(* Logix 5000 project; controller MV vendor 1 type 14 code 217 rev 31.11; software revision 31.00; part 5 of 53 *)
(* tags used below, declared in another part *)
   Always_Off : BOOL;
   Always_On : BOOL;
   ChangeDayONS : BOOL;
   CheckTimeMask : INT;
   CLOCKsetvalues : DINT[7];
   CurrentTime : DateTime;
   CWD : CHECKWORD_FLAGS;
   FtoF_raw_input : REAL;
   ItoF_raw_input : INT;
   MC_ALARM_RETURNED_STRING : STRING;
   MC_CH1_Log_ID : DINT;
   MC_CH2_Log_ID : DINT;
   MC_Channel1_Channel_1_event : STRING;
   MC_Channel1_Channel_1_event_prefix : STRING;
   MC_Channel1_Channel_2_event : STRING;
   MC_Channel1_Channel_2_event_prefix : STRING;
   MC_CLOCK_system_set : BOOL;
   MC_DetTank1_Service_event : STRING;
   MC_DetTank1_Service_event_prefix : STRING;
   MC_DetTank2_Service_event : STRING;
   MC_DetTank2_Service_event_prefix : STRING;
   MC_Event_Alarm_Tag : ALARM_DIGITAL;
   MC_Event_control_FIFO : CONTROL;
   MC_Event_control_FIFO_Operation_Type : CONTROL;
   MC_Event_Delay_For_Data : TIMER;
   MC_Event_Delay_For_PLC_Startup_Data : TIMER;
   MC_Event_Delay_Timer : TIMER;
   MC_Event_Delay_Timer_Off : TIMER;
   MC_Event_from_buffer : STRING;
   MC_Event_from_buffer_LogData1 : REAL;
   MC_Event_from_buffer_LogData2 : REAL;
   MC_Event_from_buffer_LogData3 : REAL;
   MC_Event_from_buffer_LogData4 : REAL;
   MC_Event_from_buffer_Operation_Type : DINT;
   MC_event_step : DINT;
   MC_Event_String_Last : STRING;
   MC_Event_Transact_Trigger_Tag : DINT;
   MC_Events_FIFO_Buffer : STRING[31];
   MC_Events_FIFO_Buffer_Operation_Type : INT[31];
   MC_Last_LogData_For_Op : REAL[60,20];
   MC_N10 : INT[255];   // SETTINGS
   MC_N100 : INT[255];   // C1_PLC Channel 1 PLC data
   MC_N100_20_alarm : ALARM_DIGITAL;
   MC_N100_20_Alarm_Ready : BOOL;
   MC_N100_20_Delayed_Timer2 : TIMER;
   MC_N100_20_Fault_Returned : STRING;
   MC_N100_20_SQL_Done : DINT;
   MC_N100_23_alarm : ALARM_DIGITAL;
   MC_N100_23_Alarm_Ready : BOOL;
   MC_N100_23_Delayed_Timer2 : TIMER;
   MC_N100_23_Event_Returned : STRING;
   MC_N100_23_SQL_Done : DINT;
   MC_N120 : INT[255];   // C2 PLC Channel 2 PLC data
   MC_N120_20_alarm : ALARM_DIGITAL;
   MC_N120_20_Alarm_Ready : BOOL;
   MC_N120_20_Delayed_Timer2 : TIMER;
   MC_N120_20_Fault_Returned : STRING;
   MC_N120_20_SQL_Done : DINT;
   MC_N120_23_alarm : ALARM_DIGITAL;
   MC_N120_23_Alarm_Ready : BOOL;
   MC_N120_23_Delayed_Timer2 : TIMER;
   MC_N120_23_Event_Returned : STRING;
   MC_N120_23_SQL_Done : DINT;
   MC_N140 : INT[31];   // RT FILL RT filling routine d ata
   MC_N160 : INT[255];   // P40 CHECK
   MC_N80 : INT[255];   // SRV1_PLC Detergent tank 1 ser vice PLC data
   MC_N80_10_alarm : ALARM_DIGITAL;
   MC_N80_10_Alarm_Ready : BOOL;
   MC_N80_10_Delayed_Timer2 : TIMER;
   MC_N80_10_Fault_Returned : STRING;
   MC_N80_10_SQL_Done : DINT;
   MC_N80_13_alarm : ALARM_DIGITAL;
   MC_N80_13_Alarm_Ready : BOOL;
   MC_N80_13_Delayed_Timer2 : TIMER;
   MC_N80_13_Event_Returned : STRING;
   MC_N80_13_SQL_Done : DINT;
   MC_N90 : INT[255];   // SV2_PLC Detergent tank 2 ser vice PLC data
   MC_N90_10_alarm : ALARM_DIGITAL;
   MC_N90_10_Alarm_Ready : BOOL;
   MC_N90_10_Delayed_Timer2 : TIMER;
   MC_N90_10_Fault_Returned : STRING;
   MC_N90_10_SQL_Done : DINT;
   MC_N90_13_alarm : ALARM_DIGITAL;
   MC_N90_13_Alarm_Ready : BOOL;
   MC_N90_13_Delayed_Timer2 : TIMER;
   MC_N90_13_Event_Returned : STRING;
   MC_N90_13_SQL_Done : DINT;
   MC_RT_Emptying_Log_ID : DINT;
   MC_RT_Filling_Log_ID : DINT;
   MC_SFile : INT[255];   // SLC Equivalent System File, So Original Code Can Remain
   MC_SRV1_Log_ID : DINT;
   MC_SRV2_Log_ID : DINT;
   One_Minute_One_Scan : BOOL;
   One_Minute_One_Scan_Timer : TIMER;
   One_Second_1_scan : BOOL;
   One_Second_One_Scan : ALIAS FOR One_Second_1_scan;
   scada_watchdog : DINT;
   scale_analog_int : DINT;
   scale_analog_result : REAL;
   scale_eu_max : REAL;
   scale_eu_min : REAL;
   scale_raw_input : REAL;
   scale_raw_max : REAL;
   scale_raw_min : REAL;
   scale_routine_active : BOOL;
   scale_temp : REAL;
(* MC_Common, continued *)

ROUTINE Analog_scale_ftof   (* ladder *)
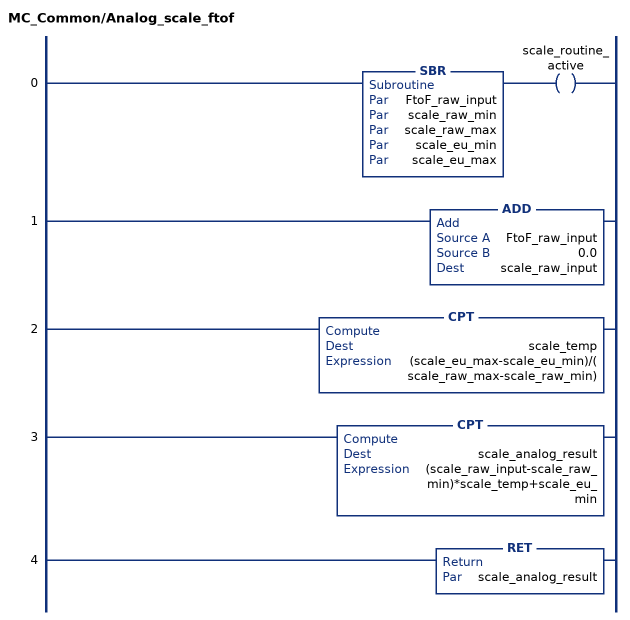
   0: SBR(FtoF_raw_input,scale_raw_min,scale_raw_max,scale_eu_min,scale_eu_max)OTE(scale_routine_active);
   1: ADD(FtoF_raw_input,0.0,scale_raw_input);
   2: CPT(scale_temp,(scale_eu_max-scale_eu_min)/(scale_raw_max-scale_raw_min));
   3: CPT(scale_analog_result,(scale_raw_input-scale_raw_min)*scale_temp+scale_eu_min);
   4: RET(scale_analog_result);
END_ROUTINE

ROUTINE Analog_Scale_FtoI   (* ladder *)
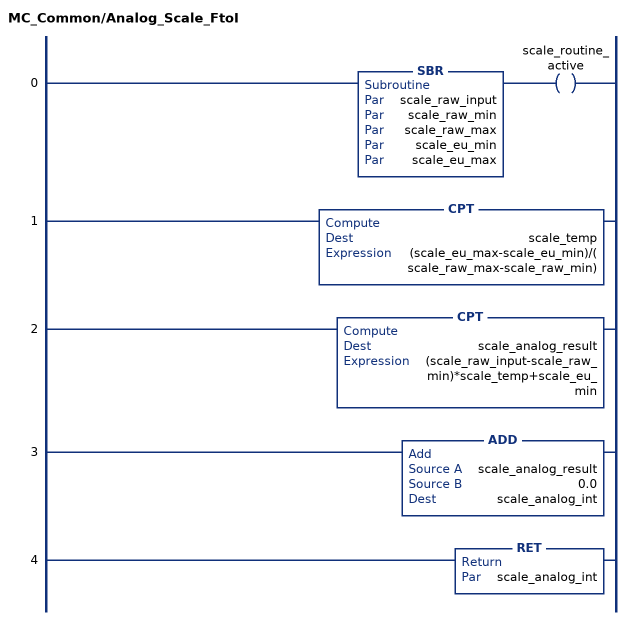
   0: SBR(scale_raw_input,scale_raw_min,scale_raw_max,scale_eu_min,scale_eu_max)OTE(scale_routine_active);
   1: CPT(scale_temp,(scale_eu_max-scale_eu_min)/(scale_raw_max-scale_raw_min));
   2: CPT(scale_analog_result,(scale_raw_input-scale_raw_min)*scale_temp+scale_eu_min);
   3: ADD(scale_analog_result,0.0,scale_analog_int);
   4: RET(scale_analog_int);
END_ROUTINE

ROUTINE Analog_Scale_ItoF   (* ladder *)
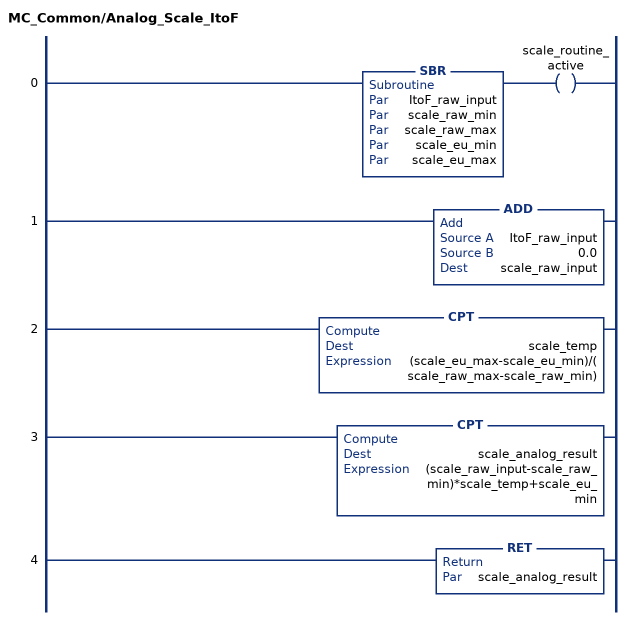
   0: SBR(ItoF_raw_input,scale_raw_min,scale_raw_max,scale_eu_min,scale_eu_max)OTE(scale_routine_active);
   1: ADD(ItoF_raw_input,0.0,scale_raw_input);
   2: CPT(scale_temp,(scale_eu_max-scale_eu_min)/(scale_raw_max-scale_raw_min));
   3: CPT(scale_analog_result,(scale_raw_input-scale_raw_min)*scale_temp+scale_eu_min);
   4: RET(scale_analog_result);
END_ROUTINE

ROUTINE ClockRoutines   (* ladder *)
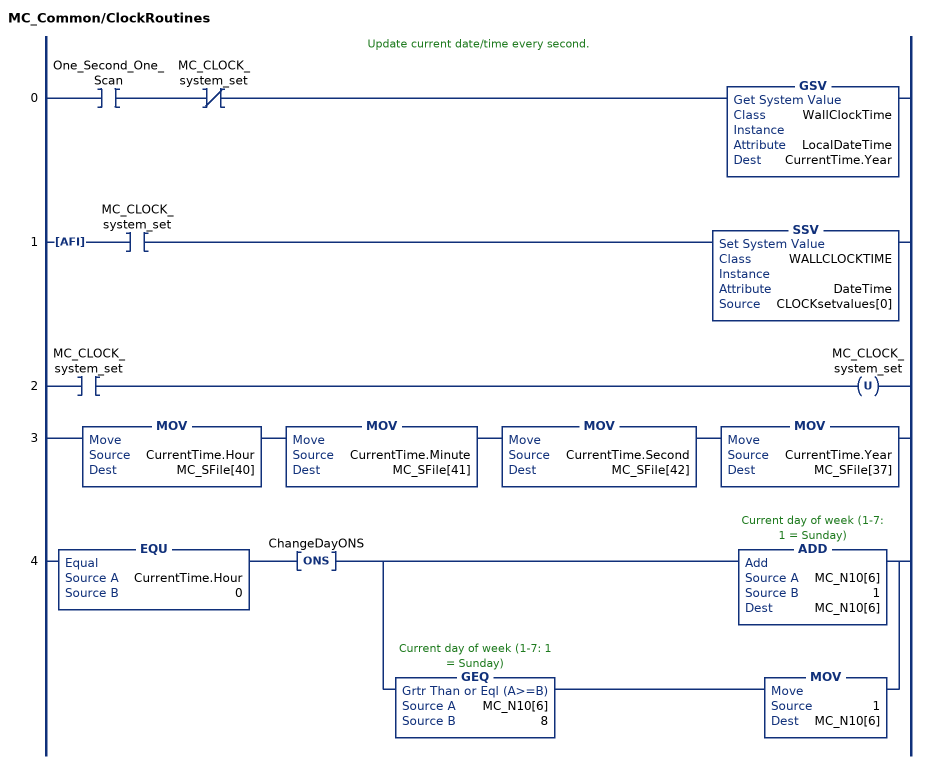
   // Update current date/time every second.
   0: XIC(One_Second_One_Scan)XIO(MC_CLOCK_system_set)GSV(WallClockTime,,LocalDateTime,CurrentTime.Year);
   1: AFI()XIC(MC_CLOCK_system_set)SSV(WALLCLOCKTIME,,DateTime,CLOCKsetvalues[0]);
   2: XIC(MC_CLOCK_system_set)OTU(MC_CLOCK_system_set);
   3: MOV(CurrentTime.Hour,MC_SFile[40])MOV(CurrentTime.Minute,MC_SFile[41])MOV(CurrentTime.Second,MC_SFile[42])MOV(CurrentTime.Year,MC_SFile[37]);
   4: EQU(CurrentTime.Hour,0)ONS(ChangeDayONS)[ADD(MC_N10[6],1,MC_N10[6]) ,GEQ(MC_N10[6],8) MOV(1,MC_N10[6]) ];
END_ROUTINE

ROUTINE Constants   (* ladder *)
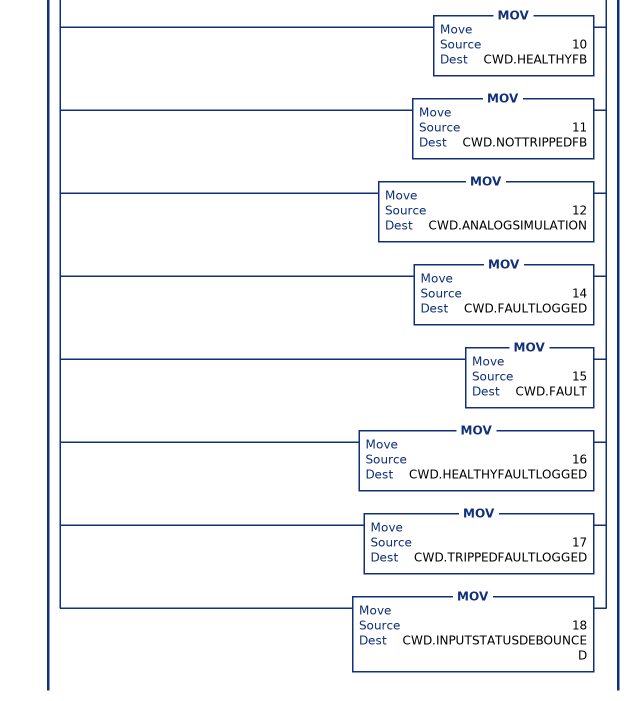
   0: [MOV(0,CWD.AUTODRV) ,MOV(0,CWD.INPUTSTATUS) ,MOV(1,CWD.PREVSCAN) ,MOV(2,CWD.SIMFAIL) ,MOV(3,CWD.OPENFB) ,MOV(3,CWD.RUNFB) ,MOV(4,CWD.CLOSEDFB) ,MOV(5,CWD.MANDRV) ,MOV(6,CWD.MANUAL) ,MOV(7,CWD.OUTPUT) ,MOV(8,CWD.CHECKOFF) ,MOV(9,CWD.HIGHLIGHT) ,MOV(10,CWD.HEALTHYFB) ,MOV(11,CWD.NOTTRIPPEDFB) ,MOV(12,CWD.ANALOGSIMULATION) ,MOV(14,CWD.FAULTLOGGED) ,MOV(15,CWD.FAULT) ,MOV(16,CWD.HEALTHYFAULTLOGGED) ,MOV(17,CWD.TRIPPEDFAULTLOGGED) ,MOV(18,CWD.INPUTSTATUSDEBOUNCED) ];
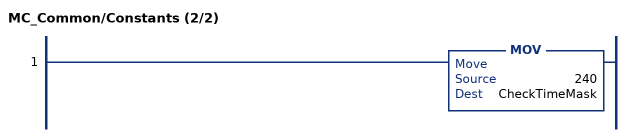
   1: MOV(240,CheckTimeMask);
END_ROUTINE

ROUTINE general_timers   (* ladder *)
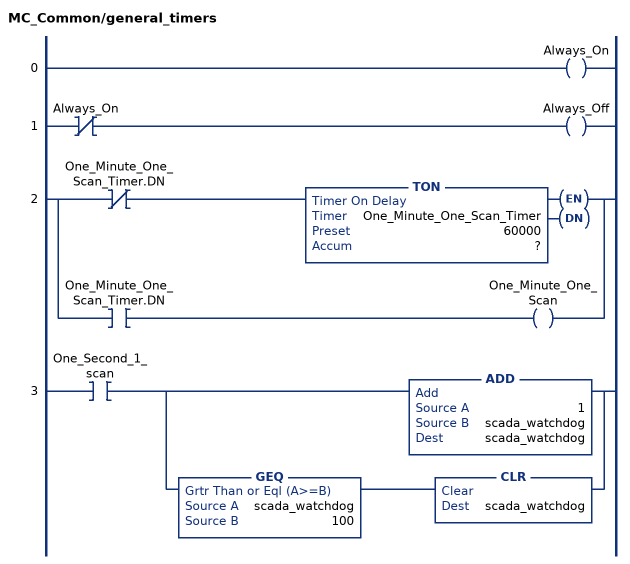
   0: OTE(Always_On);
   1: XIO(Always_On)OTE(Always_Off);
   2: [XIO(One_Minute_One_Scan_Timer.DN) TON(One_Minute_One_Scan_Timer,?,?) ,XIC(One_Minute_One_Scan_Timer.DN) OTE(One_Minute_One_Scan) ];
   3: XIC(One_Second_1_scan)[ADD(1,scada_watchdog,scada_watchdog) ,GEQ(scada_watchdog,100) CLR(scada_watchdog) ];
END_ROUTINE

ROUTINE MC_A_Alarms_From_PLC   (* ladder *)
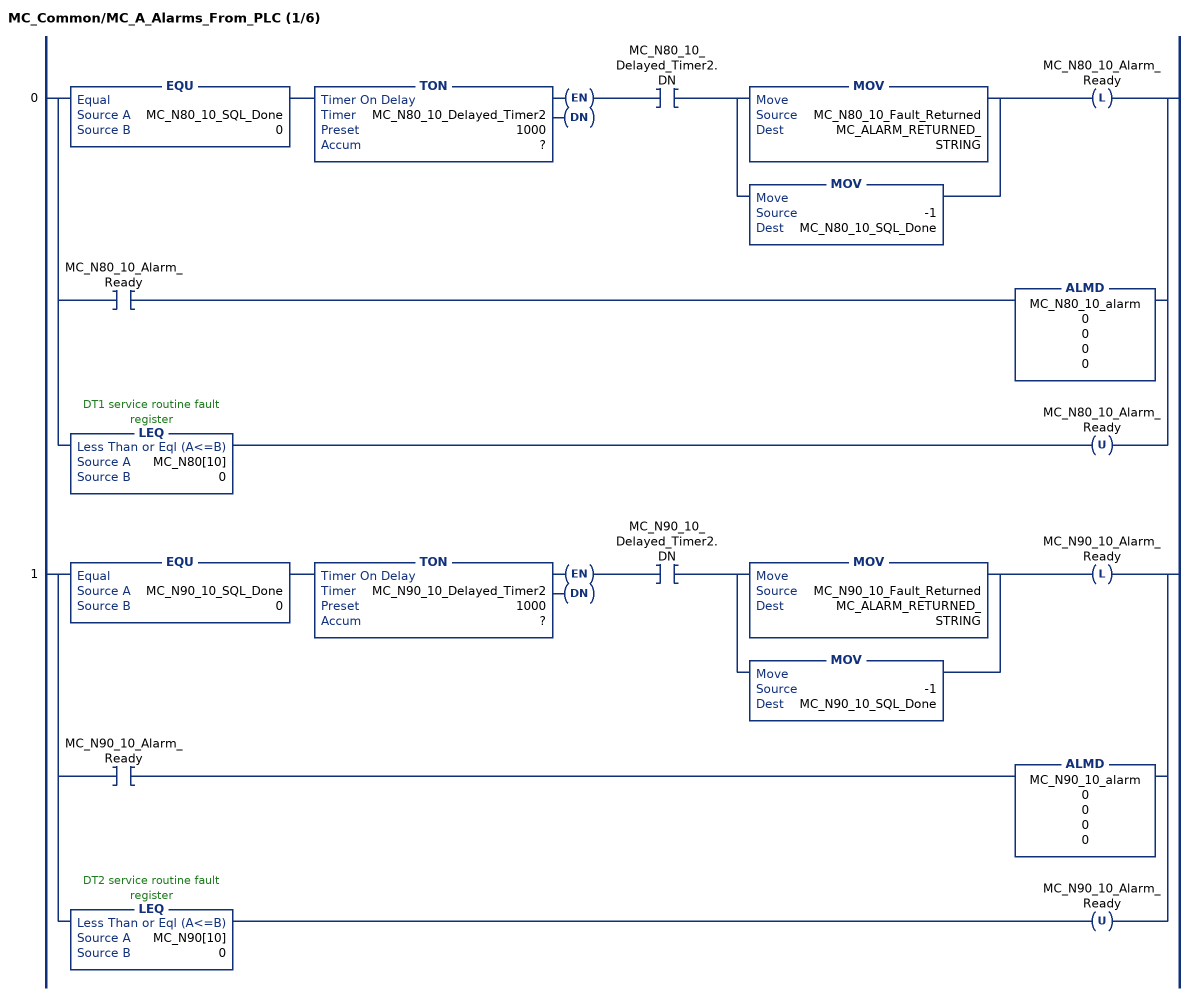
   0: [EQU(MC_N80_10_SQL_Done,0) TON(MC_N80_10_Delayed_Timer2,?,?) XIC(MC_N80_10_Delayed_Timer2.DN) [MOV(MC_N80_10_Fault_Returned,MC_ALARM_RETURNED_STRING) ,MOV(-1,MC_N80_10_SQL_Done) ] OTL(MC_N80_10_Alarm_Ready) ,XIC(MC_N80_10_Alarm_Ready) ALMD(MC_N80_10_alarm,0,0,0,0) ,LEQ(MC_N80[10],0) OTU(MC_N80_10_Alarm_Ready) ];
   1: [EQU(MC_N90_10_SQL_Done,0) TON(MC_N90_10_Delayed_Timer2,?,?) XIC(MC_N90_10_Delayed_Timer2.DN) [MOV(MC_N90_10_Fault_Returned,MC_ALARM_RETURNED_STRING) ,MOV(-1,MC_N90_10_SQL_Done) ] OTL(MC_N90_10_Alarm_Ready) ,XIC(MC_N90_10_Alarm_Ready) ALMD(MC_N90_10_alarm,0,0,0,0) ,LEQ(MC_N90[10],0) OTU(MC_N90_10_Alarm_Ready) ];
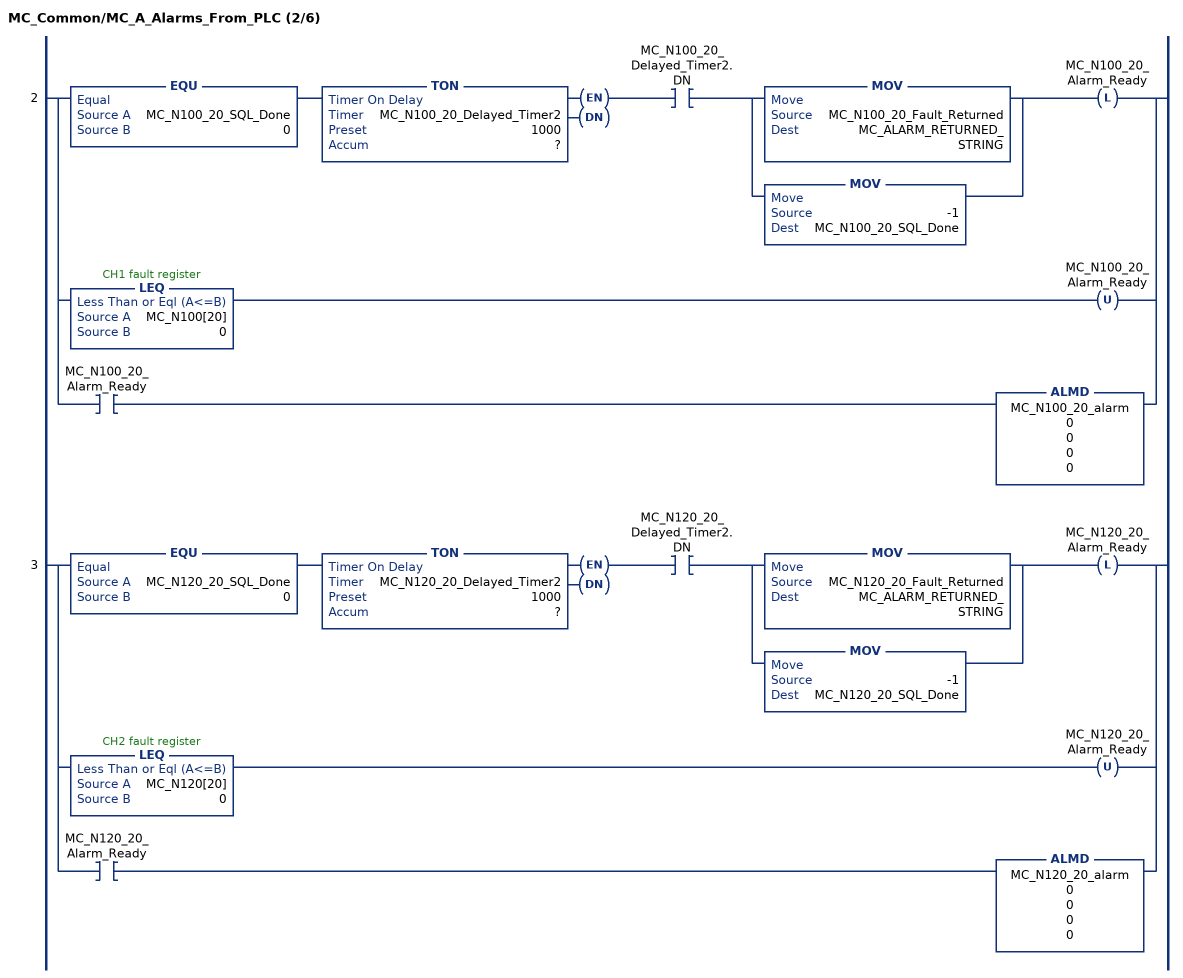
   2: [EQU(MC_N100_20_SQL_Done,0) TON(MC_N100_20_Delayed_Timer2,?,?) XIC(MC_N100_20_Delayed_Timer2.DN) [MOV(MC_N100_20_Fault_Returned,MC_ALARM_RETURNED_STRING) ,MOV(-1,MC_N100_20_SQL_Done) ] OTL(MC_N100_20_Alarm_Ready) ,LEQ(MC_N100[20],0) OTU(MC_N100_20_Alarm_Ready) ,XIC(MC_N100_20_Alarm_Ready) ALMD(MC_N100_20_alarm,0,0,0,0) ];
   3: [EQU(MC_N120_20_SQL_Done,0) TON(MC_N120_20_Delayed_Timer2,?,?) XIC(MC_N120_20_Delayed_Timer2.DN) [MOV(MC_N120_20_Fault_Returned,MC_ALARM_RETURNED_STRING) ,MOV(-1,MC_N120_20_SQL_Done) ] OTL(MC_N120_20_Alarm_Ready) ,LEQ(MC_N120[20],0) OTU(MC_N120_20_Alarm_Ready) ,XIC(MC_N120_20_Alarm_Ready) ALMD(MC_N120_20_alarm,0,0,0,0) ];
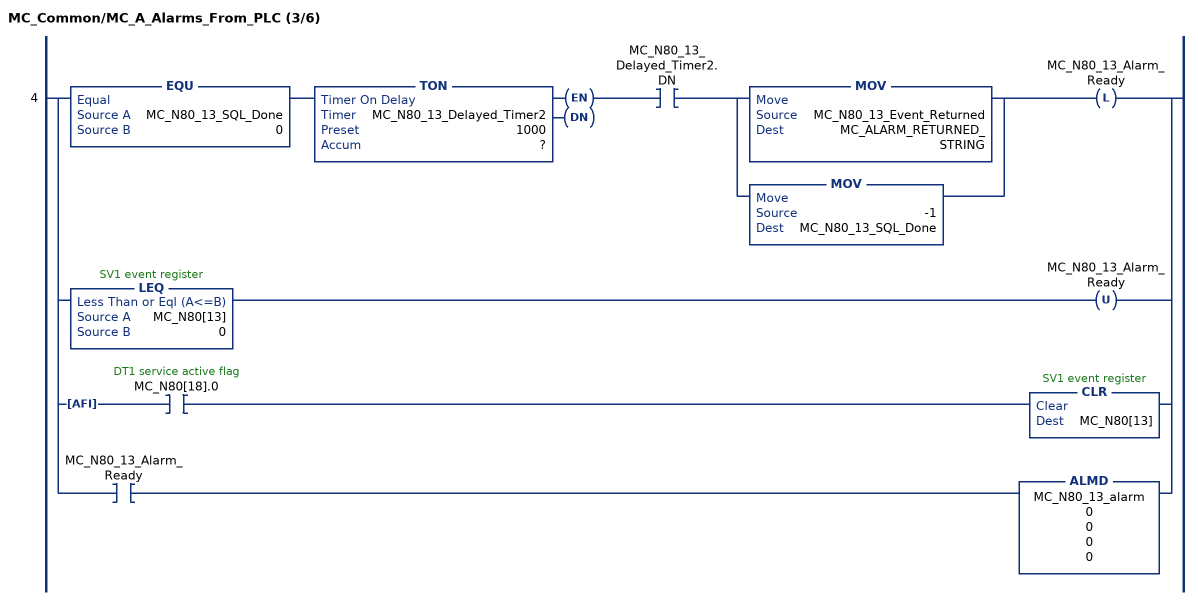
   4: [EQU(MC_N80_13_SQL_Done,0) TON(MC_N80_13_Delayed_Timer2,?,?) XIC(MC_N80_13_Delayed_Timer2.DN) [MOV(MC_N80_13_Event_Returned,MC_ALARM_RETURNED_STRING) ,MOV(-1,MC_N80_13_SQL_Done) ] OTL(MC_N80_13_Alarm_Ready) ,LEQ(MC_N80[13],0) OTU(MC_N80_13_Alarm_Ready) ,AFI() XIC(MC_N80[18].0) CLR(MC_N80[13]) ,XIC(MC_N80_13_Alarm_Ready) ALMD(MC_N80_13_alarm,0,0,0,0) ];
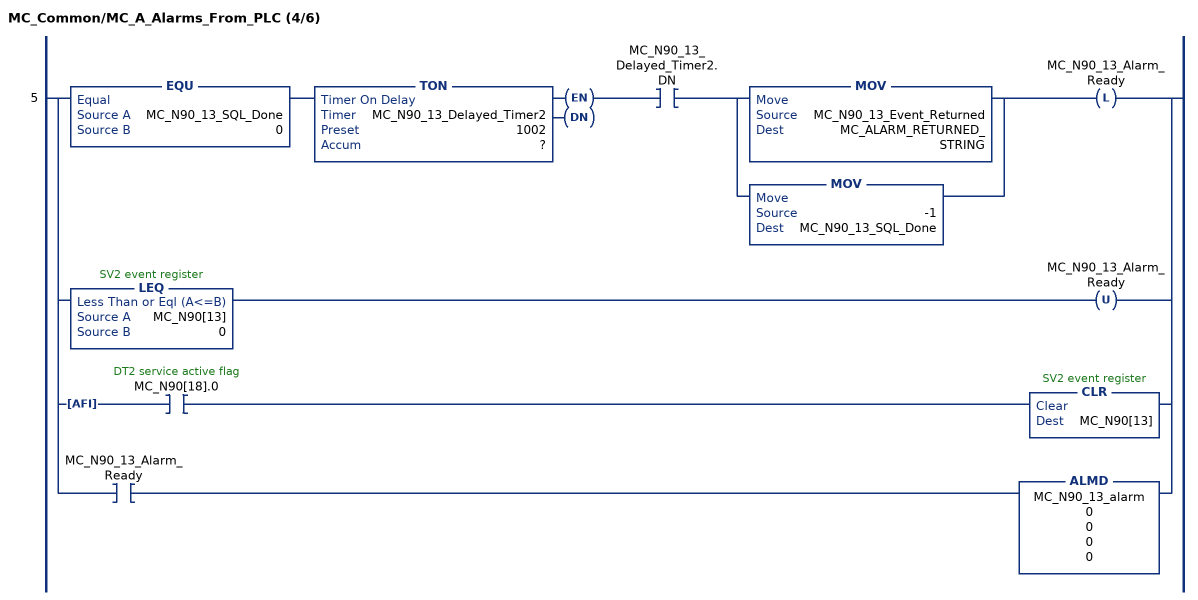
   5: [EQU(MC_N90_13_SQL_Done,0) TON(MC_N90_13_Delayed_Timer2,?,?) XIC(MC_N90_13_Delayed_Timer2.DN) [MOV(MC_N90_13_Event_Returned,MC_ALARM_RETURNED_STRING) ,MOV(-1,MC_N90_13_SQL_Done) ] OTL(MC_N90_13_Alarm_Ready) ,LEQ(MC_N90[13],0) OTU(MC_N90_13_Alarm_Ready) ,AFI() XIC(MC_N90[18].0) CLR(MC_N90[13]) ,XIC(MC_N90_13_Alarm_Ready) ALMD(MC_N90_13_alarm,0,0,0,0) ];
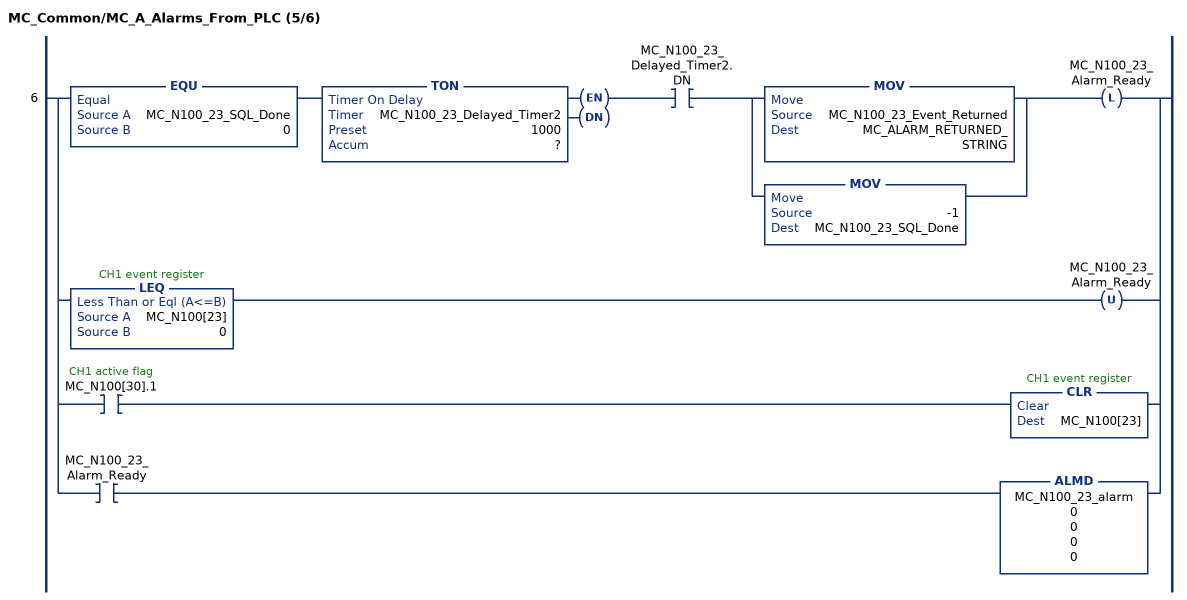
   6: [EQU(MC_N100_23_SQL_Done,0) TON(MC_N100_23_Delayed_Timer2,?,?) XIC(MC_N100_23_Delayed_Timer2.DN) [MOV(MC_N100_23_Event_Returned,MC_ALARM_RETURNED_STRING) ,MOV(-1,MC_N100_23_SQL_Done) ] OTL(MC_N100_23_Alarm_Ready) ,LEQ(MC_N100[23],0) OTU(MC_N100_23_Alarm_Ready) ,XIC(MC_N100[30].1) CLR(MC_N100[23]) ,XIC(MC_N100_23_Alarm_Ready) ALMD(MC_N100_23_alarm,0,0,0,0) ];
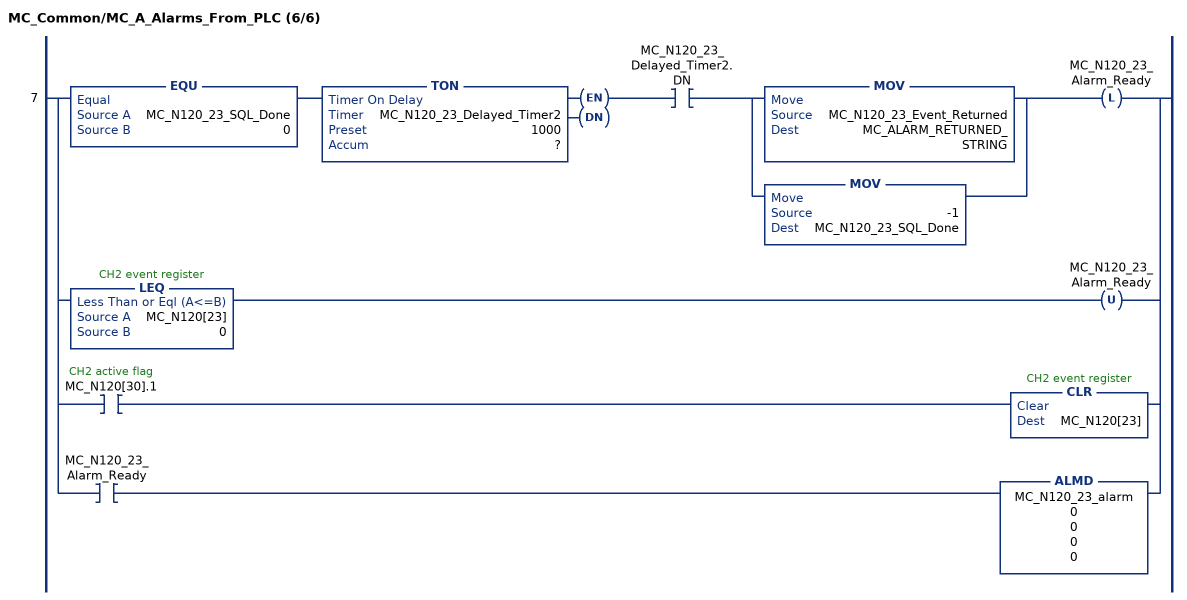
   7: [EQU(MC_N120_23_SQL_Done,0) TON(MC_N120_23_Delayed_Timer2,?,?) XIC(MC_N120_23_Delayed_Timer2.DN) [MOV(MC_N120_23_Event_Returned,MC_ALARM_RETURNED_STRING) ,MOV(-1,MC_N120_23_SQL_Done) ] OTL(MC_N120_23_Alarm_Ready) ,LEQ(MC_N120[23],0) OTU(MC_N120_23_Alarm_Ready) ,XIC(MC_N120[30].1) CLR(MC_N120[23]) ,XIC(MC_N120_23_Alarm_Ready) ALMD(MC_N120_23_alarm,0,0,0,0) ];
END_ROUTINE

ROUTINE MC_A_Events_From_Scada   (* ladder *)
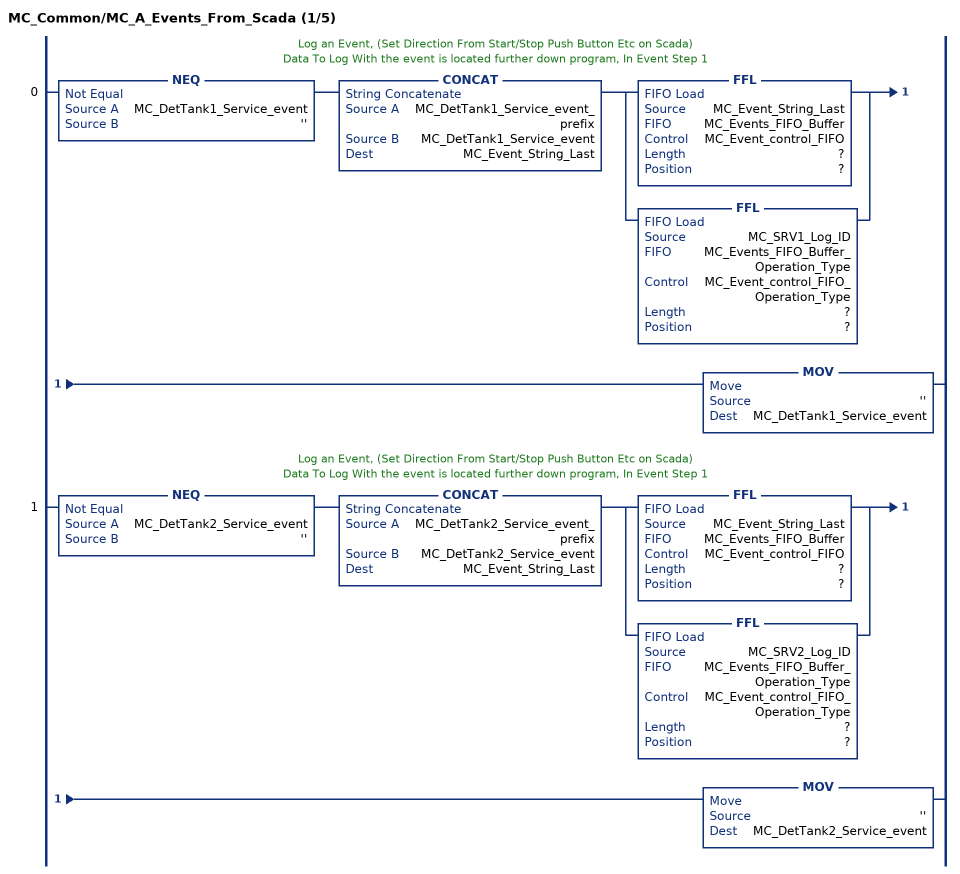
   // Log an Event, (Set Direction From Start/Stop Push Button Etc on Scada)
   // Data To Log With the event is located further down program, In Event Step 1
   0: NEQ(MC_DetTank1_Service_event,'')CONCAT(MC_DetTank1_Service_event_prefix,MC_DetTank1_Service_event,MC_Event_String_Last)[FFL(MC_Event_String_Last,MC_Events_FIFO_Buffer,MC_Event_control_FIFO,?,?) ,FFL(MC_SRV1_Log_ID,MC_Events_FIFO_Buffer_Operation_Type,MC_Event_control_FIFO_Operation_Type,?,?) ]MOV('',MC_DetTank1_Service_event);
   // Log an Event, (Set Direction From Start/Stop Push Button Etc on Scada)
   // Data To Log With the event is located further down program, In Event Step 1
   1: NEQ(MC_DetTank2_Service_event,'')CONCAT(MC_DetTank2_Service_event_prefix,MC_DetTank2_Service_event,MC_Event_String_Last)[FFL(MC_Event_String_Last,MC_Events_FIFO_Buffer,MC_Event_control_FIFO,?,?) ,FFL(MC_SRV2_Log_ID,MC_Events_FIFO_Buffer_Operation_Type,MC_Event_control_FIFO_Operation_Type,?,?) ]MOV('',MC_DetTank2_Service_event);
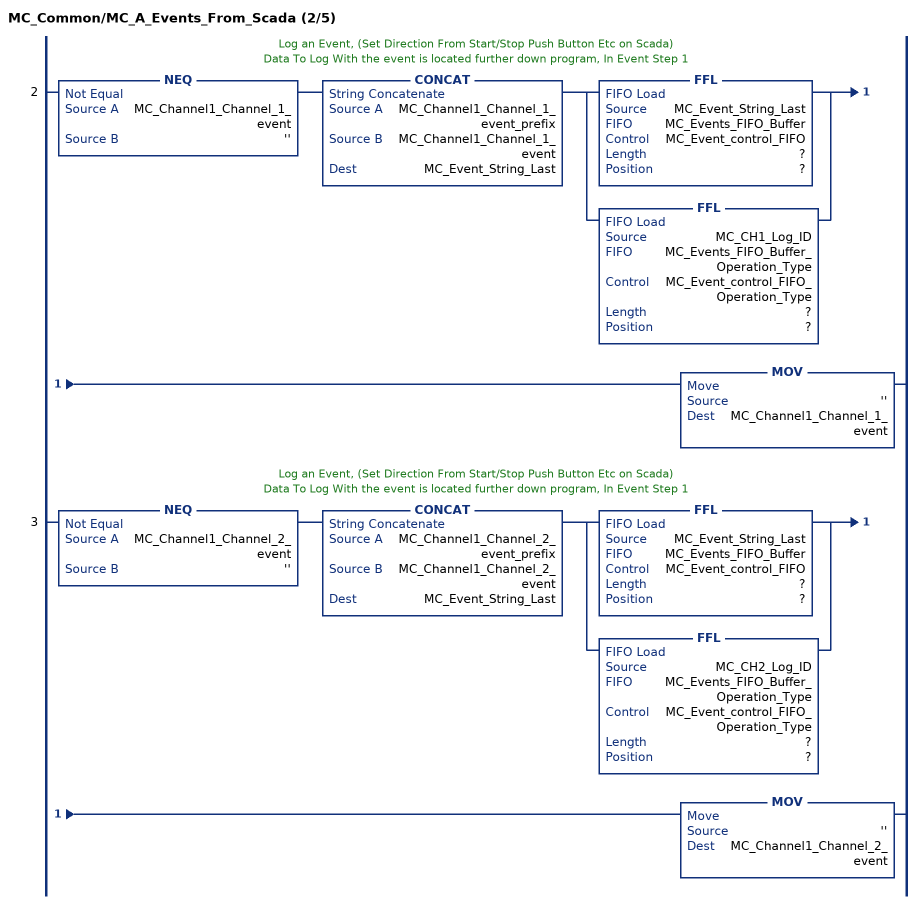
   // Log an Event, (Set Direction From Start/Stop Push Button Etc on Scada)
   // Data To Log With the event is located further down program, In Event Step 1
   2: NEQ(MC_Channel1_Channel_1_event,'')CONCAT(MC_Channel1_Channel_1_event_prefix,MC_Channel1_Channel_1_event,MC_Event_String_Last)[FFL(MC_Event_String_Last,MC_Events_FIFO_Buffer,MC_Event_control_FIFO,?,?) ,FFL(MC_CH1_Log_ID,MC_Events_FIFO_Buffer_Operation_Type,MC_Event_control_FIFO_Operation_Type,?,?) ]MOV('',MC_Channel1_Channel_1_event);
   // Log an Event, (Set Direction From Start/Stop Push Button Etc on Scada)
   // Data To Log With the event is located further down program, In Event Step 1
   3: NEQ(MC_Channel1_Channel_2_event,'')CONCAT(MC_Channel1_Channel_2_event_prefix,MC_Channel1_Channel_2_event,MC_Event_String_Last)[FFL(MC_Event_String_Last,MC_Events_FIFO_Buffer,MC_Event_control_FIFO,?,?) ,FFL(MC_CH2_Log_ID,MC_Events_FIFO_Buffer_Operation_Type,MC_Event_control_FIFO_Operation_Type,?,?) ]MOV('',MC_Channel1_Channel_2_event);
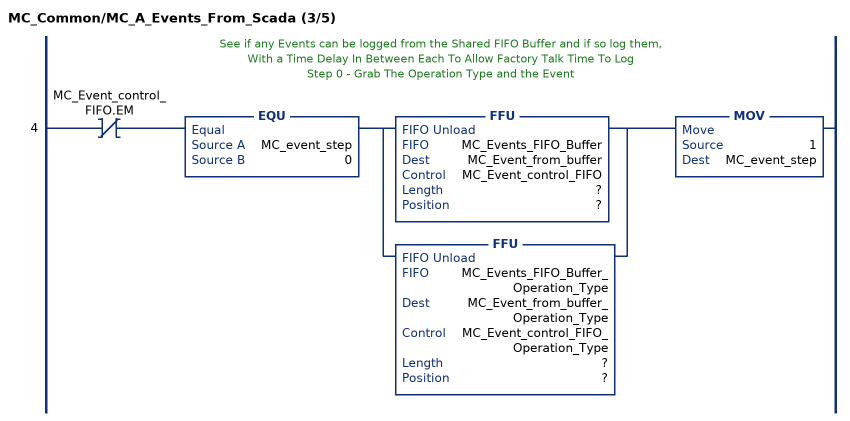
   // See if any Events can be logged from the Shared FIFO Buffer and if so log them,
   // With a Time Delay In Between Each To Allow Factory Talk Time To Log
   // Step 0 - Grab The Operation Type and the Event
   4: XIO(MC_Event_control_FIFO.EM)EQU(MC_event_step,0)[FFU(MC_Events_FIFO_Buffer,MC_Event_from_buffer,MC_Event_control_FIFO,?,?) ,FFU(MC_Events_FIFO_Buffer_Operation_Type,MC_Event_from_buffer_Operation_Type,MC_Event_control_FIFO_Operation_Type,?,?) ]MOV(1,MC_event_step);
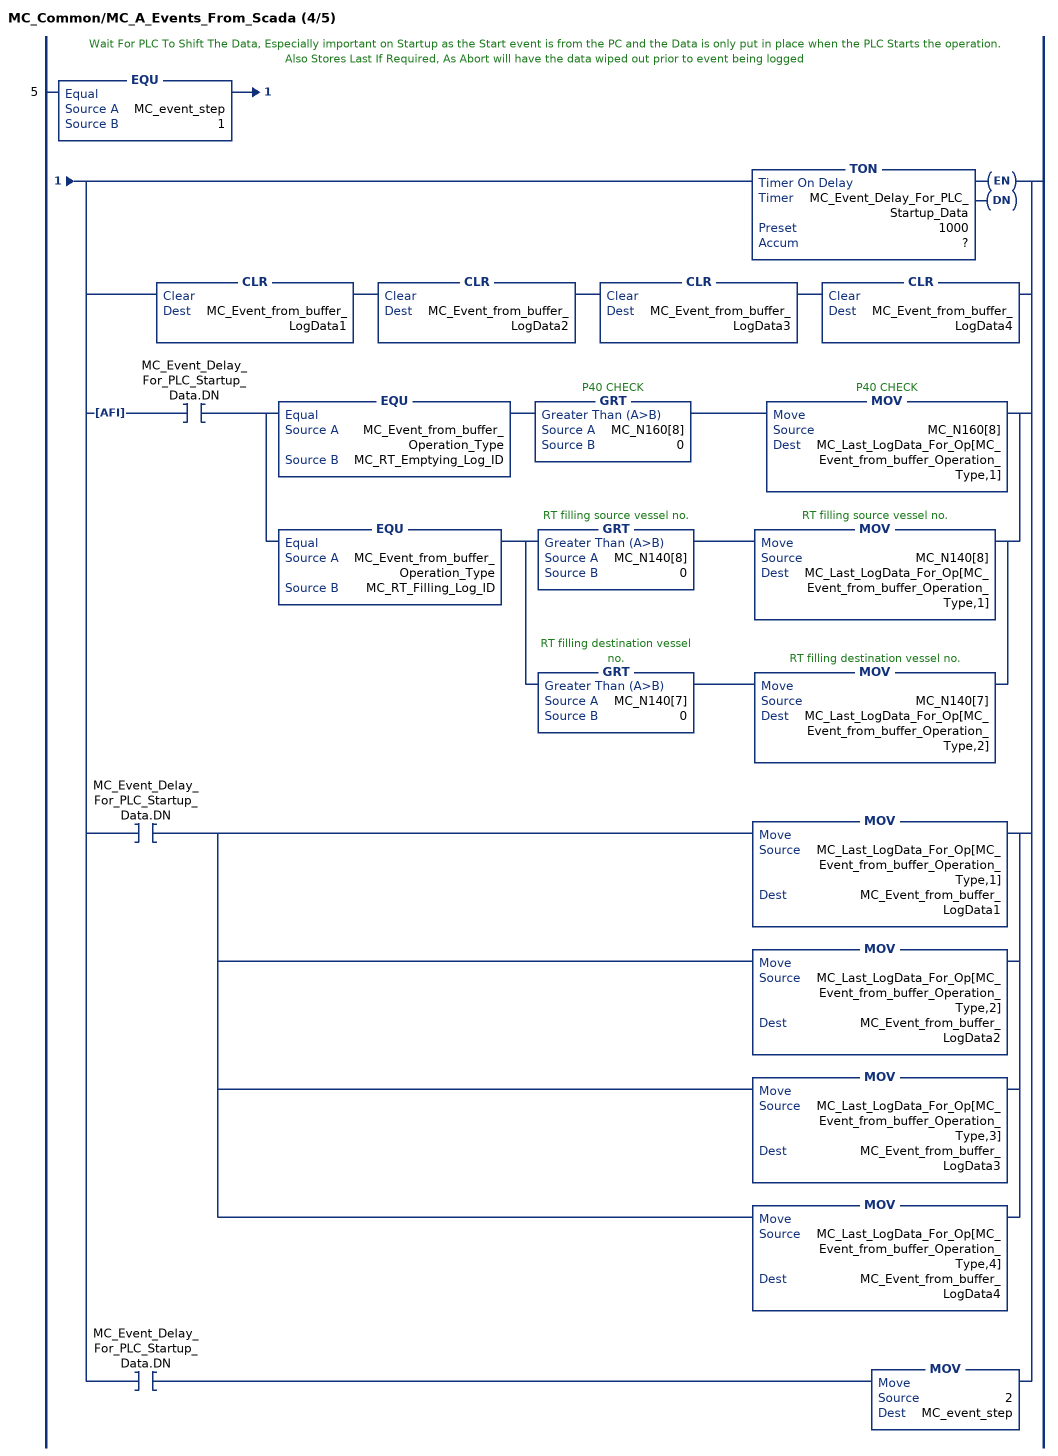
   // Wait For PLC To Shift The Data, Especially important on Startup as the Start event is from the PC and the Data is only put in place when the PLC Starts the operation.
   // Also Stores Last If Required, As Abort will have the data wiped out prior to event being logged
   5: EQU(MC_event_step,1)[TON(MC_Event_Delay_For_PLC_Startup_Data,?,?) ,CLR(MC_Event_from_buffer_LogData1) CLR(MC_Event_from_buffer_LogData2) CLR(MC_Event_from_buffer_LogData3) CLR(MC_Event_from_buffer_LogData4) ,AFI() XIC(MC_Event_Delay_For_PLC_Startup_Data.DN) [EQU(MC_Event_from_buffer_Operation_Type,MC_RT_Emptying_Log_ID) GRT(MC_N160[8],0) MOV(MC_N160[8],MC_Last_LogData_For_Op[MC_Event_from_buffer_Operation_Type,1]) ,EQU(MC_Event_from_buffer_Operation_Type,MC_RT_Filling_Log_ID) [GRT(MC_N140[8],0) MOV(MC_N140[8],MC_Last_LogData_For_Op[MC_Event_from_buffer_Operation_Type,1]) ,GRT(MC_N140[7],0) MOV(MC_N140[7],MC_Last_LogData_For_Op[MC_Event_from_buffer_Operation_Type,2]) ] ] ,XIC(MC_Event_Delay_For_PLC_Startup_Data.DN) [MOV(MC_Last_LogData_For_Op[MC_Event_from_buffer_Operation_Type,1],MC_Event_from_buffer_LogData1) ,MOV(MC_Last_LogData_For_Op[MC_Event_from_buffer_Operation_Type,2],MC_Event_from_buffer_LogData2) ,MOV(MC_Last_LogData_For_Op[MC_Event_from_buffer_Operation_Type,3],MC_Event_from_buffer_LogData3) ,MOV(MC_Last_LogData_For_Op[MC_Event_from_buffer_Operation_Type,4],MC_Event_from_buffer_LogData4) ] ,XIC(MC_Event_Delay_For_PLC_Startup_Data.DN) MOV(2,MC_event_step) ];
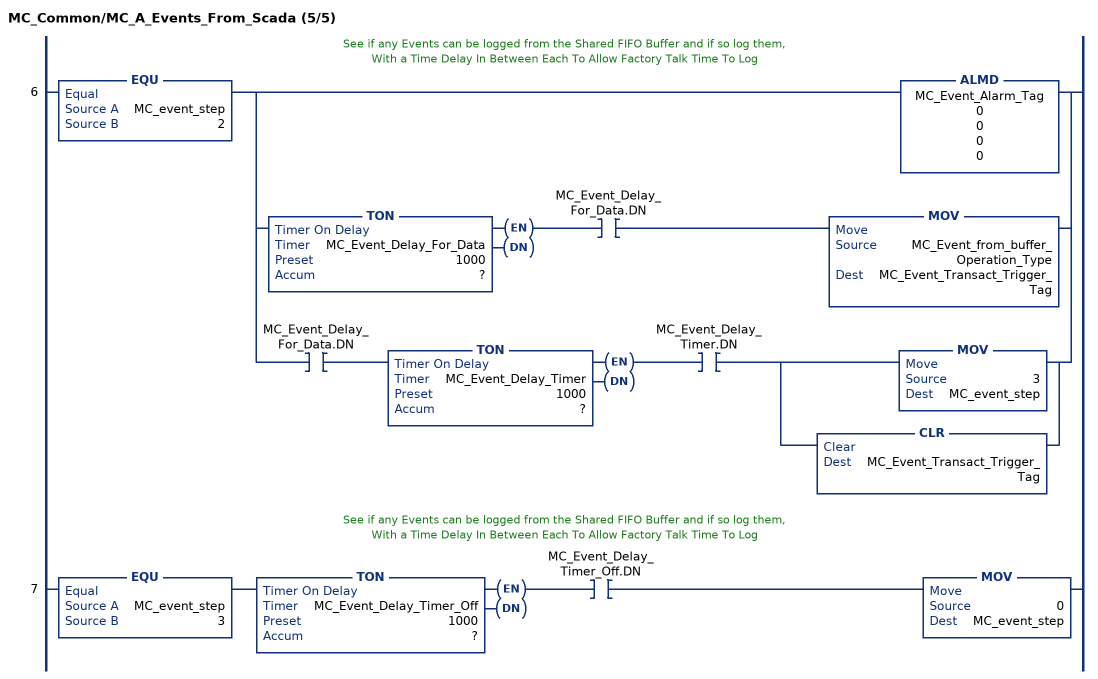
   // See if any Events can be logged from the Shared FIFO Buffer and if so log them,
   // With a Time Delay In Between Each To Allow Factory Talk Time To Log
   6: EQU(MC_event_step,2)[ALMD(MC_Event_Alarm_Tag,0,0,0,0) ,TON(MC_Event_Delay_For_Data,?,?) XIC(MC_Event_Delay_For_Data.DN) MOV(MC_Event_from_buffer_Operation_Type,MC_Event_Transact_Trigger_Tag) ,XIC(MC_Event_Delay_For_Data.DN) TON(MC_Event_Delay_Timer,?,?) XIC(MC_Event_Delay_Timer.DN) [MOV(3,MC_event_step) ,CLR(MC_Event_Transact_Trigger_Tag) ] ];
   // See if any Events can be logged from the Shared FIFO Buffer and if so log them,
   // With a Time Delay In Between Each To Allow Factory Talk Time To Log
   7: EQU(MC_event_step,3)TON(MC_Event_Delay_Timer_Off,?,?)XIC(MC_Event_Delay_Timer_Off.DN)MOV(0,MC_event_step);
END_ROUTINE
